REGION Network 145
   Label( C76_Comm_Fault )
   RUNG wire#powerrail
      Coil( "SectionComment" )
   END_RUNG
   // the same network as SCL:
   C76_Comm_Fault:
   "SectionComment" := TRUE;
END_REGION

REGION Network 146
   // **********************************************************************************************************************
   // 
   // Carrier 77 I-Device Data Transfer Interlocks from Carrier to SDC
   // 
   // **********************************************************************************************************************
   RUNG wire#powerrail
      Coil( "SectionComment" )
   END_RUNG
   // the same network as SCL:
   "SectionComment" := TRUE;
END_REGION

REGION Network 147
   RUNG wire#powerrail
      Contact( "Carrier_77_Status.0" )
      Coil( "EMS".Carrier[77].SDC_IN.HeartBeat )
   END_RUNG
   // the same network as SCL:
   "EMS".Carrier[77].SDC_IN.HeartBeat := "Carrier_77_Status.0";
END_REGION

REGION Network 148
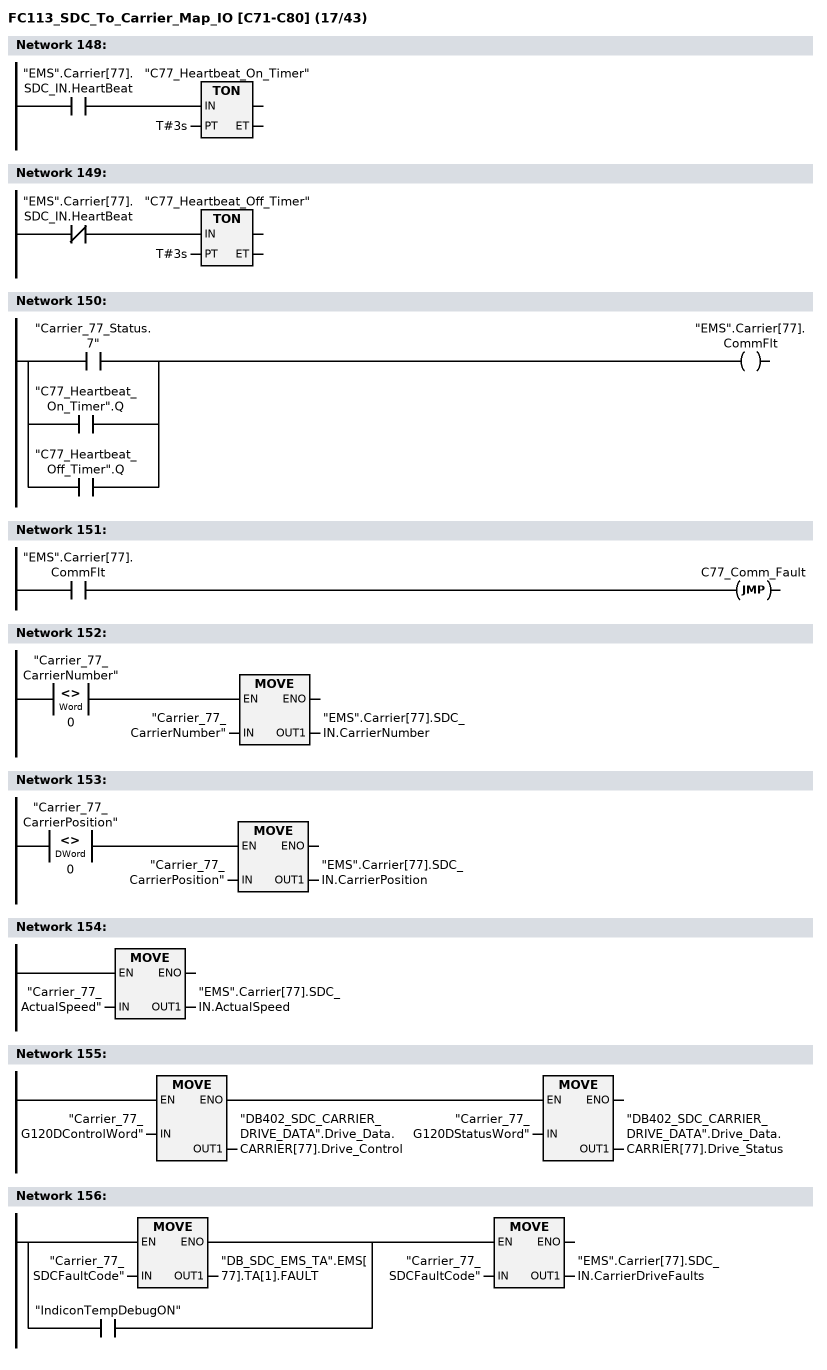
   "C77_Heartbeat_On_Timer".TON(IN := "EMS".Carrier[77].SDC_IN.HeartBeat, PT := T#3s);
END_REGION

REGION Network 149
   "C77_Heartbeat_Off_Timer".TON(IN := NOT "EMS".Carrier[77].SDC_IN.HeartBeat, PT := T#3s);
END_REGION

REGION Network 150
   RUNG wire#powerrail
      Contact( "Carrier_77_Status.7" )
      wire#w1
      Coil( "EMS".Carrier[77].CommFlt )
   END_RUNG
   RUNG wire#powerrail
      Contact( "C77_Heartbeat_On_Timer".Q )
   END_RUNG wire#w1
   RUNG wire#powerrail
      Contact( "C77_Heartbeat_Off_Timer".Q )
   END_RUNG wire#w1
   // the same network as SCL:
   "EMS".Carrier[77].CommFlt := "Carrier_77_Status.7" OR "C77_Heartbeat_On_Timer".Q OR "C77_Heartbeat_Off_Timer".Q;
END_REGION

REGION Network 151
   RUNG wire#powerrail
      Contact( "EMS".Carrier[77].CommFlt )
      JumpCoil( C77_Comm_Fault )
   END_RUNG
   // the same network as SCL:
   IF "EMS".Carrier[77].CommFlt THEN GOTO C77_Comm_Fault; END_IF;
END_REGION

REGION Network 152
   RUNG wire#powerrail
      { S7_Templates := "SrcType := Word" } NE_Contact(in1 := "Carrier_77_CarrierNumber", in2 := 0)
      Move(in := "Carrier_77_CarrierNumber", out1 => "EMS".Carrier[77].SDC_IN.CarrierNumber)
   END_RUNG
   // the same network as SCL:
   IF "Carrier_77_CarrierNumber" <> 0 THEN
       "EMS".Carrier[77].SDC_IN.CarrierNumber := "Carrier_77_CarrierNumber";
   END_IF;
END_REGION

REGION Network 153
   RUNG wire#powerrail
      { S7_Templates := "SrcType := DWord" } NE_Contact(in1 := "Carrier_77_CarrierPosition", in2 := 0)
      Move(in := "Carrier_77_CarrierPosition", out1 => "EMS".Carrier[77].SDC_IN.CarrierPosition)
   END_RUNG
   // the same network as SCL:
   IF "Carrier_77_CarrierPosition" <> 0 THEN
       "EMS".Carrier[77].SDC_IN.CarrierPosition := "Carrier_77_CarrierPosition";
   END_IF;
END_REGION

REGION Network 154
   RUNG wire#powerrail
      Move(in := "Carrier_77_ActualSpeed", out1 => "EMS".Carrier[77].SDC_IN.ActualSpeed)
   END_RUNG
   // the same network as SCL:
   "EMS".Carrier[77].SDC_IN.ActualSpeed := "Carrier_77_ActualSpeed";
END_REGION

REGION Network 155
   RUNG wire#powerrail
      Move(in := "Carrier_77_G120DControlWord", out1 => "DB402_SDC_CARRIER_DRIVE_DATA".Drive_Data.CARRIER[77].Drive_Control)
      Move(in := "Carrier_77_G120DStatusWord", out1 => "DB402_SDC_CARRIER_DRIVE_DATA".Drive_Data.CARRIER[77].Drive_Status)
   END_RUNG
   // the same network as SCL:
   "DB402_SDC_CARRIER_DRIVE_DATA".Drive_Data.CARRIER[77].Drive_Control := "Carrier_77_G120DControlWord";
   "DB402_SDC_CARRIER_DRIVE_DATA".Drive_Data.CARRIER[77].Drive_Status := "Carrier_77_G120DStatusWord";
END_REGION

REGION Network 156
   RUNG wire#powerrail
      Move(in := "Carrier_77_SDCFaultCode", out1 => "DB_SDC_EMS_TA".EMS[77].TA[1].FAULT)
      wire#w1
      Move(in := "Carrier_77_SDCFaultCode", out1 => "EMS".Carrier[77].SDC_IN.CarrierDriveFaults)
   END_RUNG
   RUNG wire#powerrail
      Contact( "IndiconTempDebugON" )
   END_RUNG wire#w1
   // the same network as SCL:
   "DB_SDC_EMS_TA".EMS[77].TA[1].FAULT := "Carrier_77_SDCFaultCode";
   IF TRUE OR "IndiconTempDebugON" THEN
       "EMS".Carrier[77].SDC_IN.CarrierDriveFaults := "Carrier_77_SDCFaultCode";
   END_IF;
END_REGION

REGION Network 157
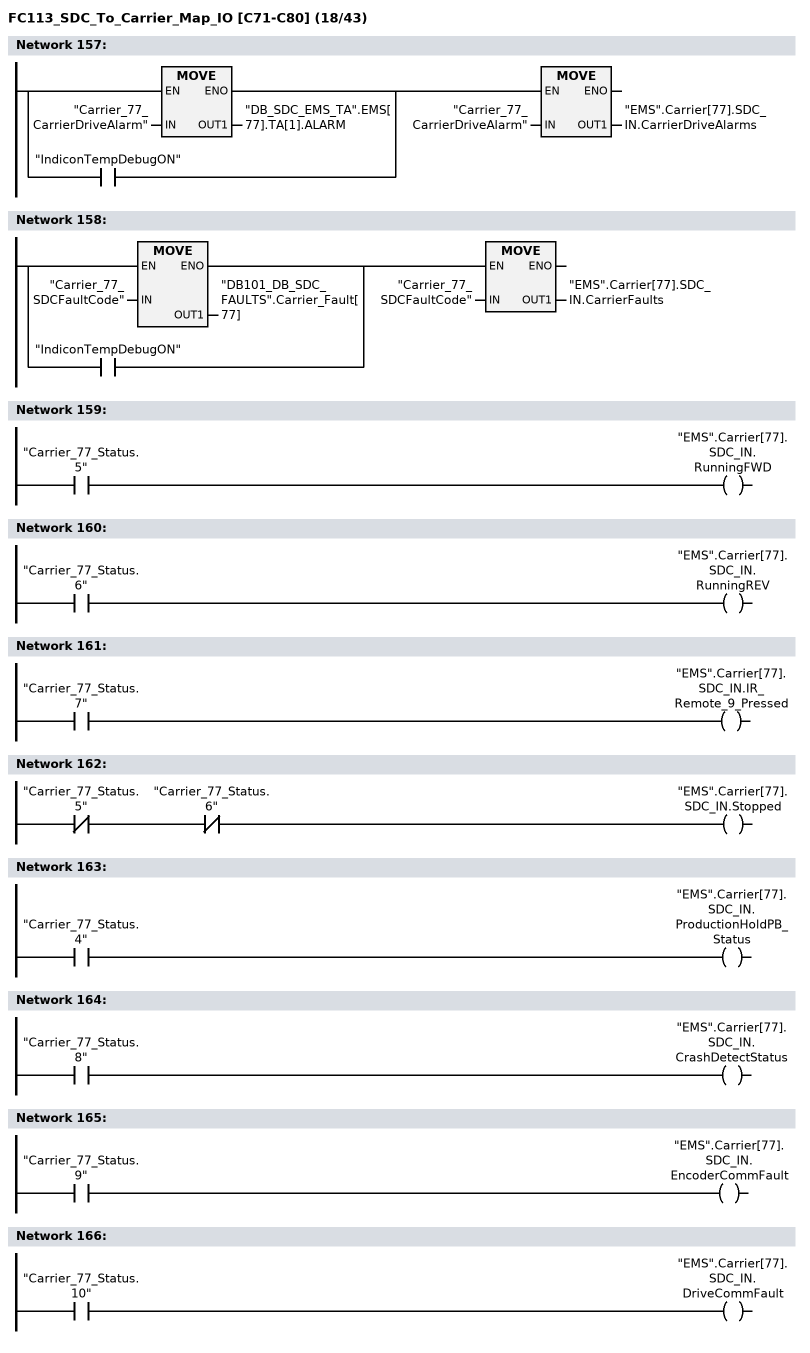
   RUNG wire#powerrail
      Move(in := "Carrier_77_CarrierDriveAlarm", out1 => "DB_SDC_EMS_TA".EMS[77].TA[1].ALARM)
      wire#w1
      Move(in := "Carrier_77_CarrierDriveAlarm", out1 => "EMS".Carrier[77].SDC_IN.CarrierDriveAlarms)
   END_RUNG
   RUNG wire#powerrail
      Contact( "IndiconTempDebugON" )
   END_RUNG wire#w1
   // the same network as SCL:
   "DB_SDC_EMS_TA".EMS[77].TA[1].ALARM := "Carrier_77_CarrierDriveAlarm";
   IF TRUE OR "IndiconTempDebugON" THEN
       "EMS".Carrier[77].SDC_IN.CarrierDriveAlarms := "Carrier_77_CarrierDriveAlarm";
   END_IF;
END_REGION

REGION Network 158
   RUNG wire#powerrail
      Move(in := "Carrier_77_SDCFaultCode", out1 => "DB101_DB_SDC_FAULTS".Carrier_Fault[77])
      wire#w1
      Move(in := "Carrier_77_SDCFaultCode", out1 => "EMS".Carrier[77].SDC_IN.CarrierFaults)
   END_RUNG
   RUNG wire#powerrail
      Contact( "IndiconTempDebugON" )
   END_RUNG wire#w1
   // the same network as SCL:
   "DB101_DB_SDC_FAULTS".Carrier_Fault[77] := "Carrier_77_SDCFaultCode";
   IF TRUE OR "IndiconTempDebugON" THEN
       "EMS".Carrier[77].SDC_IN.CarrierFaults := "Carrier_77_SDCFaultCode";
   END_IF;
END_REGION

REGION Network 159
   RUNG wire#powerrail
      Contact( "Carrier_77_Status.5" )
      Coil( "EMS".Carrier[77].SDC_IN.RunningFWD )
   END_RUNG
   // the same network as SCL:
   "EMS".Carrier[77].SDC_IN.RunningFWD := "Carrier_77_Status.5";
END_REGION

REGION Network 160
   RUNG wire#powerrail
      Contact( "Carrier_77_Status.6" )
      Coil( "EMS".Carrier[77].SDC_IN.RunningREV )
   END_RUNG
   // the same network as SCL:
   "EMS".Carrier[77].SDC_IN.RunningREV := "Carrier_77_Status.6";
END_REGION

REGION Network 161
   RUNG wire#powerrail
      Contact( "Carrier_77_Status.7" )
      Coil( "EMS".Carrier[77].SDC_IN.IR_Remote_9_Pressed )
   END_RUNG
   // the same network as SCL:
   "EMS".Carrier[77].SDC_IN.IR_Remote_9_Pressed := "Carrier_77_Status.7";
END_REGION

REGION Network 162
   RUNG wire#powerrail
      I_Contact( "Carrier_77_Status.5" )
      I_Contact( "Carrier_77_Status.6" )
      Coil( "EMS".Carrier[77].SDC_IN.Stopped )
   END_RUNG
   // the same network as SCL:
   "EMS".Carrier[77].SDC_IN.Stopped := NOT "Carrier_77_Status.5" AND NOT "Carrier_77_Status.6";
END_REGION

REGION Network 163
   RUNG wire#powerrail
      Contact( "Carrier_77_Status.4" )
      Coil( "EMS".Carrier[77].SDC_IN.ProductionHoldPB_Status )
   END_RUNG
   // the same network as SCL:
   "EMS".Carrier[77].SDC_IN.ProductionHoldPB_Status := "Carrier_77_Status.4";
END_REGION

REGION Network 164
   RUNG wire#powerrail
      Contact( "Carrier_77_Status.8" )
      Coil( "EMS".Carrier[77].SDC_IN.CrashDetectStatus )
   END_RUNG
   // the same network as SCL:
   "EMS".Carrier[77].SDC_IN.CrashDetectStatus := "Carrier_77_Status.8";
END_REGION

REGION Network 165
   RUNG wire#powerrail
      Contact( "Carrier_77_Status.9" )
      Coil( "EMS".Carrier[77].SDC_IN.EncoderCommFault )
   END_RUNG
   // the same network as SCL:
   "EMS".Carrier[77].SDC_IN.EncoderCommFault := "Carrier_77_Status.9";
END_REGION

REGION Network 166
   RUNG wire#powerrail
      Contact( "Carrier_77_Status.10" )
      Coil( "EMS".Carrier[77].SDC_IN.DriveCommFault )
   END_RUNG
   // the same network as SCL:
   "EMS".Carrier[77].SDC_IN.DriveCommFault := "Carrier_77_Status.10";
END_REGION

REGION Network 167
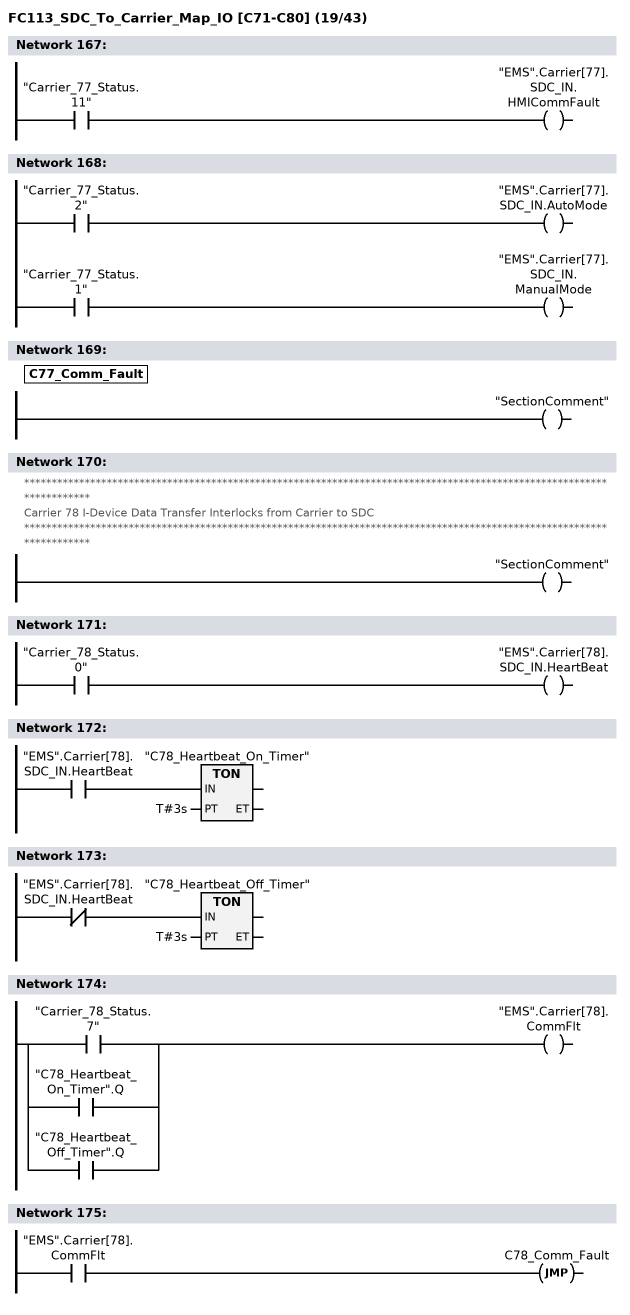
   RUNG wire#powerrail
      Contact( "Carrier_77_Status.11" )
      Coil( "EMS".Carrier[77].SDC_IN.HMICommFault )
   END_RUNG
   // the same network as SCL:
   "EMS".Carrier[77].SDC_IN.HMICommFault := "Carrier_77_Status.11";
END_REGION

REGION Network 168
   RUNG wire#powerrail
      Contact( "Carrier_77_Status.2" )
      Coil( "EMS".Carrier[77].SDC_IN.AutoMode )
   END_RUNG
   RUNG wire#powerrail
      Contact( "Carrier_77_Status.1" )
      Coil( "EMS".Carrier[77].SDC_IN.ManualMode )
   END_RUNG
   // the same network as SCL:
   "EMS".Carrier[77].SDC_IN.AutoMode := "Carrier_77_Status.2";
   "EMS".Carrier[77].SDC_IN.ManualMode := "Carrier_77_Status.1";
END_REGION

REGION Network 169
   Label( C77_Comm_Fault )
   RUNG wire#powerrail
      Coil( "SectionComment" )
   END_RUNG
   // the same network as SCL:
   C77_Comm_Fault:
   "SectionComment" := TRUE;
END_REGION

REGION Network 170
   // **********************************************************************************************************************
   // 
   // Carrier 78 I-Device Data Transfer Interlocks from Carrier to SDC
   // 
   // **********************************************************************************************************************
   RUNG wire#powerrail
      Coil( "SectionComment" )
   END_RUNG
   // the same network as SCL:
   "SectionComment" := TRUE;
END_REGION

REGION Network 171
   RUNG wire#powerrail
      Contact( "Carrier_78_Status.0" )
      Coil( "EMS".Carrier[78].SDC_IN.HeartBeat )
   END_RUNG
   // the same network as SCL:
   "EMS".Carrier[78].SDC_IN.HeartBeat := "Carrier_78_Status.0";
END_REGION

REGION Network 172
   "C78_Heartbeat_On_Timer".TON(IN := "EMS".Carrier[78].SDC_IN.HeartBeat, PT := T#3s);
END_REGION

REGION Network 173
   "C78_Heartbeat_Off_Timer".TON(IN := NOT "EMS".Carrier[78].SDC_IN.HeartBeat, PT := T#3s);
END_REGION

REGION Network 174
   RUNG wire#powerrail
      Contact( "Carrier_78_Status.7" )
      wire#w1
      Coil( "EMS".Carrier[78].CommFlt )
   END_RUNG
   RUNG wire#powerrail
      Contact( "C78_Heartbeat_On_Timer".Q )
   END_RUNG wire#w1
   RUNG wire#powerrail
      Contact( "C78_Heartbeat_Off_Timer".Q )
   END_RUNG wire#w1
   // the same network as SCL:
   "EMS".Carrier[78].CommFlt := "Carrier_78_Status.7" OR "C78_Heartbeat_On_Timer".Q OR "C78_Heartbeat_Off_Timer".Q;
END_REGION

REGION Network 175
   RUNG wire#powerrail
      Contact( "EMS".Carrier[78].CommFlt )
      JumpCoil( C78_Comm_Fault )
   END_RUNG
   // the same network as SCL:
   IF "EMS".Carrier[78].CommFlt THEN GOTO C78_Comm_Fault; END_IF;
END_REGION

REGION Network 176
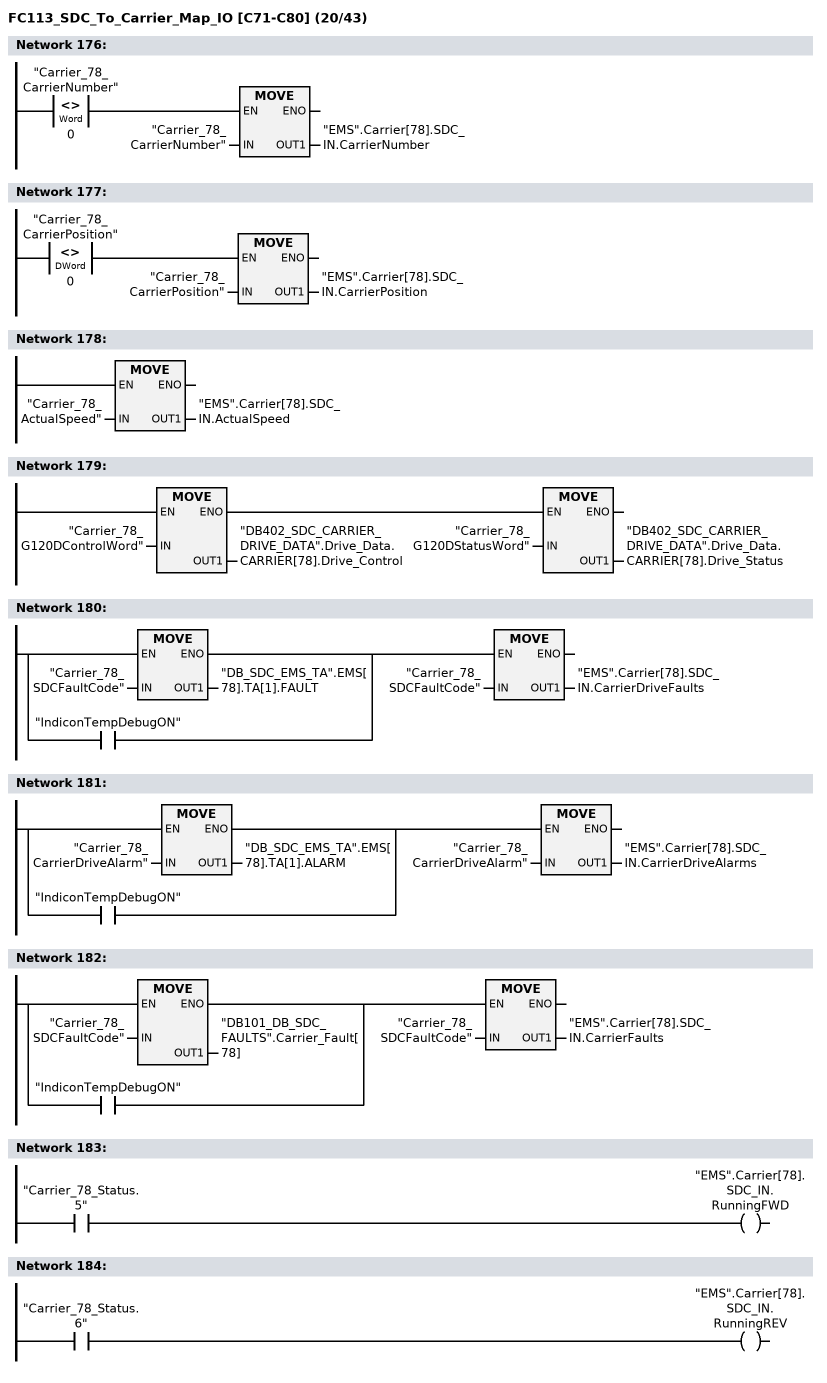
   RUNG wire#powerrail
      { S7_Templates := "SrcType := Word" } NE_Contact(in1 := "Carrier_78_CarrierNumber", in2 := 0)
      Move(in := "Carrier_78_CarrierNumber", out1 => "EMS".Carrier[78].SDC_IN.CarrierNumber)
   END_RUNG
   // the same network as SCL:
   IF "Carrier_78_CarrierNumber" <> 0 THEN
       "EMS".Carrier[78].SDC_IN.CarrierNumber := "Carrier_78_CarrierNumber";
   END_IF;
END_REGION

REGION Network 177
   RUNG wire#powerrail
      { S7_Templates := "SrcType := DWord" } NE_Contact(in1 := "Carrier_78_CarrierPosition", in2 := 0)
      Move(in := "Carrier_78_CarrierPosition", out1 => "EMS".Carrier[78].SDC_IN.CarrierPosition)
   END_RUNG
   // the same network as SCL:
   IF "Carrier_78_CarrierPosition" <> 0 THEN
       "EMS".Carrier[78].SDC_IN.CarrierPosition := "Carrier_78_CarrierPosition";
   END_IF;
END_REGION

REGION Network 178
   RUNG wire#powerrail
      Move(in := "Carrier_78_ActualSpeed", out1 => "EMS".Carrier[78].SDC_IN.ActualSpeed)
   END_RUNG
   // the same network as SCL:
   "EMS".Carrier[78].SDC_IN.ActualSpeed := "Carrier_78_ActualSpeed";
END_REGION

REGION Network 179
   RUNG wire#powerrail
      Move(in := "Carrier_78_G120DControlWord", out1 => "DB402_SDC_CARRIER_DRIVE_DATA".Drive_Data.CARRIER[78].Drive_Control)
      Move(in := "Carrier_78_G120DStatusWord", out1 => "DB402_SDC_CARRIER_DRIVE_DATA".Drive_Data.CARRIER[78].Drive_Status)
   END_RUNG
   // the same network as SCL:
   "DB402_SDC_CARRIER_DRIVE_DATA".Drive_Data.CARRIER[78].Drive_Control := "Carrier_78_G120DControlWord";
   "DB402_SDC_CARRIER_DRIVE_DATA".Drive_Data.CARRIER[78].Drive_Status := "Carrier_78_G120DStatusWord";
END_REGION

REGION Network 180
   RUNG wire#powerrail
      Move(in := "Carrier_78_SDCFaultCode", out1 => "DB_SDC_EMS_TA".EMS[78].TA[1].FAULT)
      wire#w1
      Move(in := "Carrier_78_SDCFaultCode", out1 => "EMS".Carrier[78].SDC_IN.CarrierDriveFaults)
   END_RUNG
   RUNG wire#powerrail
      Contact( "IndiconTempDebugON" )
   END_RUNG wire#w1
   // the same network as SCL:
   "DB_SDC_EMS_TA".EMS[78].TA[1].FAULT := "Carrier_78_SDCFaultCode";
   IF TRUE OR "IndiconTempDebugON" THEN
       "EMS".Carrier[78].SDC_IN.CarrierDriveFaults := "Carrier_78_SDCFaultCode";
   END_IF;
END_REGION

REGION Network 181
   RUNG wire#powerrail
      Move(in := "Carrier_78_CarrierDriveAlarm", out1 => "DB_SDC_EMS_TA".EMS[78].TA[1].ALARM)
      wire#w1
      Move(in := "Carrier_78_CarrierDriveAlarm", out1 => "EMS".Carrier[78].SDC_IN.CarrierDriveAlarms)
   END_RUNG
   RUNG wire#powerrail
      Contact( "IndiconTempDebugON" )
   END_RUNG wire#w1
   // the same network as SCL:
   "DB_SDC_EMS_TA".EMS[78].TA[1].ALARM := "Carrier_78_CarrierDriveAlarm";
   IF TRUE OR "IndiconTempDebugON" THEN
       "EMS".Carrier[78].SDC_IN.CarrierDriveAlarms := "Carrier_78_CarrierDriveAlarm";
   END_IF;
END_REGION

REGION Network 182
   RUNG wire#powerrail
      Move(in := "Carrier_78_SDCFaultCode", out1 => "DB101_DB_SDC_FAULTS".Carrier_Fault[78])
      wire#w1
      Move(in := "Carrier_78_SDCFaultCode", out1 => "EMS".Carrier[78].SDC_IN.CarrierFaults)
   END_RUNG
   RUNG wire#powerrail
      Contact( "IndiconTempDebugON" )
   END_RUNG wire#w1
   // the same network as SCL:
   "DB101_DB_SDC_FAULTS".Carrier_Fault[78] := "Carrier_78_SDCFaultCode";
   IF TRUE OR "IndiconTempDebugON" THEN
       "EMS".Carrier[78].SDC_IN.CarrierFaults := "Carrier_78_SDCFaultCode";
   END_IF;
END_REGION

REGION Network 183
   RUNG wire#powerrail
      Contact( "Carrier_78_Status.5" )
      Coil( "EMS".Carrier[78].SDC_IN.RunningFWD )
   END_RUNG
   // the same network as SCL:
   "EMS".Carrier[78].SDC_IN.RunningFWD := "Carrier_78_Status.5";
END_REGION

REGION Network 184
   RUNG wire#powerrail
      Contact( "Carrier_78_Status.6" )
      Coil( "EMS".Carrier[78].SDC_IN.RunningREV )
   END_RUNG
   // the same network as SCL:
   "EMS".Carrier[78].SDC_IN.RunningREV := "Carrier_78_Status.6";
END_REGION

REGION Network 185
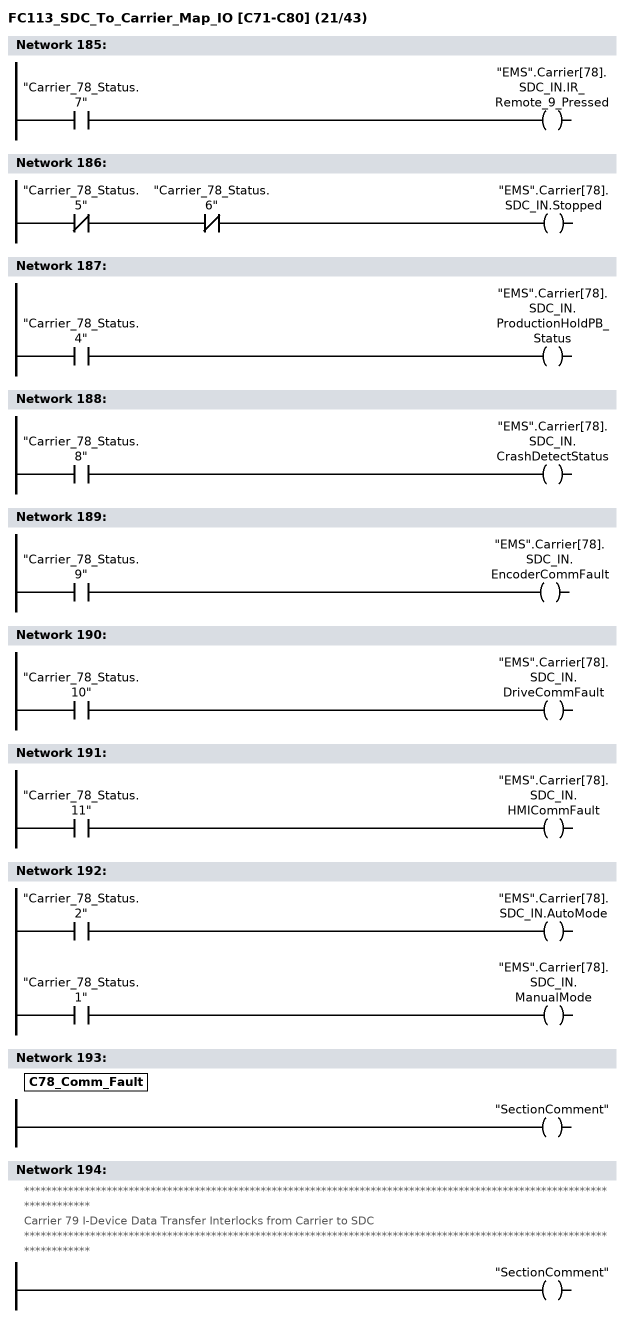
   RUNG wire#powerrail
      Contact( "Carrier_78_Status.7" )
      Coil( "EMS".Carrier[78].SDC_IN.IR_Remote_9_Pressed )
   END_RUNG
   // the same network as SCL:
   "EMS".Carrier[78].SDC_IN.IR_Remote_9_Pressed := "Carrier_78_Status.7";
END_REGION

REGION Network 186
   RUNG wire#powerrail
      I_Contact( "Carrier_78_Status.5" )
      I_Contact( "Carrier_78_Status.6" )
      Coil( "EMS".Carrier[78].SDC_IN.Stopped )
   END_RUNG
   // the same network as SCL:
   "EMS".Carrier[78].SDC_IN.Stopped := NOT "Carrier_78_Status.5" AND NOT "Carrier_78_Status.6";
END_REGION

REGION Network 187
   RUNG wire#powerrail
      Contact( "Carrier_78_Status.4" )
      Coil( "EMS".Carrier[78].SDC_IN.ProductionHoldPB_Status )
   END_RUNG
   // the same network as SCL:
   "EMS".Carrier[78].SDC_IN.ProductionHoldPB_Status := "Carrier_78_Status.4";
END_REGION

REGION Network 188
   RUNG wire#powerrail
      Contact( "Carrier_78_Status.8" )
      Coil( "EMS".Carrier[78].SDC_IN.CrashDetectStatus )
   END_RUNG
   // the same network as SCL:
   "EMS".Carrier[78].SDC_IN.CrashDetectStatus := "Carrier_78_Status.8";
END_REGION

REGION Network 189
   RUNG wire#powerrail
      Contact( "Carrier_78_Status.9" )
      Coil( "EMS".Carrier[78].SDC_IN.EncoderCommFault )
   END_RUNG
   // the same network as SCL:
   "EMS".Carrier[78].SDC_IN.EncoderCommFault := "Carrier_78_Status.9";
END_REGION

REGION Network 190
   RUNG wire#powerrail
      Contact( "Carrier_78_Status.10" )
      Coil( "EMS".Carrier[78].SDC_IN.DriveCommFault )
   END_RUNG
   // the same network as SCL:
   "EMS".Carrier[78].SDC_IN.DriveCommFault := "Carrier_78_Status.10";
END_REGION

REGION Network 191
   RUNG wire#powerrail
      Contact( "Carrier_78_Status.11" )
      Coil( "EMS".Carrier[78].SDC_IN.HMICommFault )
   END_RUNG
   // the same network as SCL:
   "EMS".Carrier[78].SDC_IN.HMICommFault := "Carrier_78_Status.11";
END_REGION

REGION Network 192
   RUNG wire#powerrail
      Contact( "Carrier_78_Status.2" )
      Coil( "EMS".Carrier[78].SDC_IN.AutoMode )
   END_RUNG
   RUNG wire#powerrail
      Contact( "Carrier_78_Status.1" )
      Coil( "EMS".Carrier[78].SDC_IN.ManualMode )
   END_RUNG
   // the same network as SCL:
   "EMS".Carrier[78].SDC_IN.AutoMode := "Carrier_78_Status.2";
   "EMS".Carrier[78].SDC_IN.ManualMode := "Carrier_78_Status.1";
END_REGION

REGION Network 193
   Label( C78_Comm_Fault )
   RUNG wire#powerrail
      Coil( "SectionComment" )
   END_RUNG
   // the same network as SCL:
   C78_Comm_Fault:
   "SectionComment" := TRUE;
END_REGION

REGION Network 194
   // **********************************************************************************************************************
   // 
   // Carrier 79 I-Device Data Transfer Interlocks from Carrier to SDC
   // 
   // **********************************************************************************************************************
   RUNG wire#powerrail
      Coil( "SectionComment" )
   END_RUNG
   // the same network as SCL:
   "SectionComment" := TRUE;
END_REGION

REGION Network 195
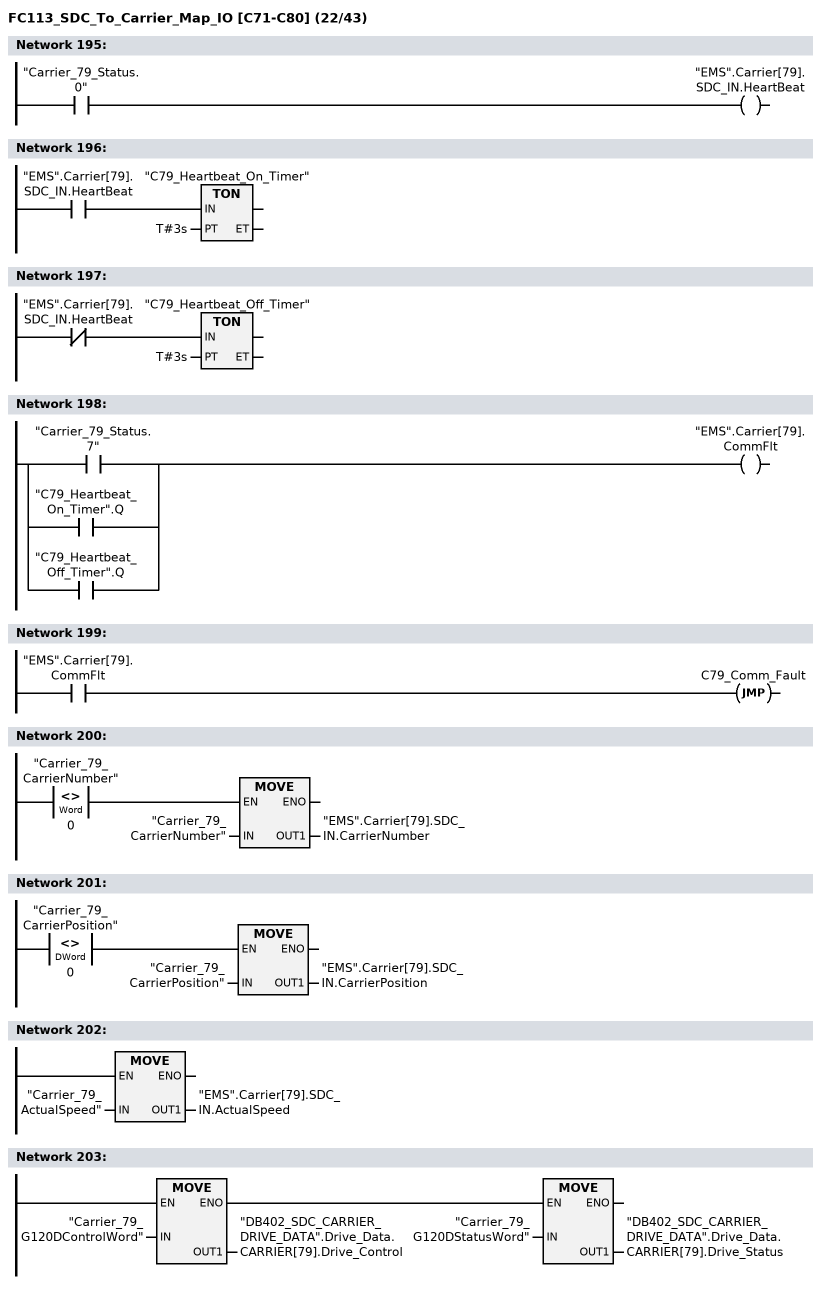
   RUNG wire#powerrail
      Contact( "Carrier_79_Status.0" )
      Coil( "EMS".Carrier[79].SDC_IN.HeartBeat )
   END_RUNG
   // the same network as SCL:
   "EMS".Carrier[79].SDC_IN.HeartBeat := "Carrier_79_Status.0";
END_REGION

REGION Network 196
   "C79_Heartbeat_On_Timer".TON(IN := "EMS".Carrier[79].SDC_IN.HeartBeat, PT := T#3s);
END_REGION

REGION Network 197
   "C79_Heartbeat_Off_Timer".TON(IN := NOT "EMS".Carrier[79].SDC_IN.HeartBeat, PT := T#3s);
END_REGION

REGION Network 198
   RUNG wire#powerrail
      Contact( "Carrier_79_Status.7" )
      wire#w1
      Coil( "EMS".Carrier[79].CommFlt )
   END_RUNG
   RUNG wire#powerrail
      Contact( "C79_Heartbeat_On_Timer".Q )
   END_RUNG wire#w1
   RUNG wire#powerrail
      Contact( "C79_Heartbeat_Off_Timer".Q )
   END_RUNG wire#w1
   // the same network as SCL:
   "EMS".Carrier[79].CommFlt := "Carrier_79_Status.7" OR "C79_Heartbeat_On_Timer".Q OR "C79_Heartbeat_Off_Timer".Q;
END_REGION

REGION Network 199
   RUNG wire#powerrail
      Contact( "EMS".Carrier[79].CommFlt )
      JumpCoil( C79_Comm_Fault )
   END_RUNG
   // the same network as SCL:
   IF "EMS".Carrier[79].CommFlt THEN GOTO C79_Comm_Fault; END_IF;
END_REGION

REGION Network 200
   RUNG wire#powerrail
      { S7_Templates := "SrcType := Word" } NE_Contact(in1 := "Carrier_79_CarrierNumber", in2 := 0)
      Move(in := "Carrier_79_CarrierNumber", out1 => "EMS".Carrier[79].SDC_IN.CarrierNumber)
   END_RUNG
   // the same network as SCL:
   IF "Carrier_79_CarrierNumber" <> 0 THEN
       "EMS".Carrier[79].SDC_IN.CarrierNumber := "Carrier_79_CarrierNumber";
   END_IF;
END_REGION

REGION Network 201
   RUNG wire#powerrail
      { S7_Templates := "SrcType := DWord" } NE_Contact(in1 := "Carrier_79_CarrierPosition", in2 := 0)
      Move(in := "Carrier_79_CarrierPosition", out1 => "EMS".Carrier[79].SDC_IN.CarrierPosition)
   END_RUNG
   // the same network as SCL:
   IF "Carrier_79_CarrierPosition" <> 0 THEN
       "EMS".Carrier[79].SDC_IN.CarrierPosition := "Carrier_79_CarrierPosition";
   END_IF;
END_REGION

REGION Network 202
   RUNG wire#powerrail
      Move(in := "Carrier_79_ActualSpeed", out1 => "EMS".Carrier[79].SDC_IN.ActualSpeed)
   END_RUNG
   // the same network as SCL:
   "EMS".Carrier[79].SDC_IN.ActualSpeed := "Carrier_79_ActualSpeed";
END_REGION

REGION Network 203
   RUNG wire#powerrail
      Move(in := "Carrier_79_G120DControlWord", out1 => "DB402_SDC_CARRIER_DRIVE_DATA".Drive_Data.CARRIER[79].Drive_Control)
      Move(in := "Carrier_79_G120DStatusWord", out1 => "DB402_SDC_CARRIER_DRIVE_DATA".Drive_Data.CARRIER[79].Drive_Status)
   END_RUNG
   // the same network as SCL:
   "DB402_SDC_CARRIER_DRIVE_DATA".Drive_Data.CARRIER[79].Drive_Control := "Carrier_79_G120DControlWord";
   "DB402_SDC_CARRIER_DRIVE_DATA".Drive_Data.CARRIER[79].Drive_Status := "Carrier_79_G120DStatusWord";
END_REGION

REGION Network 204
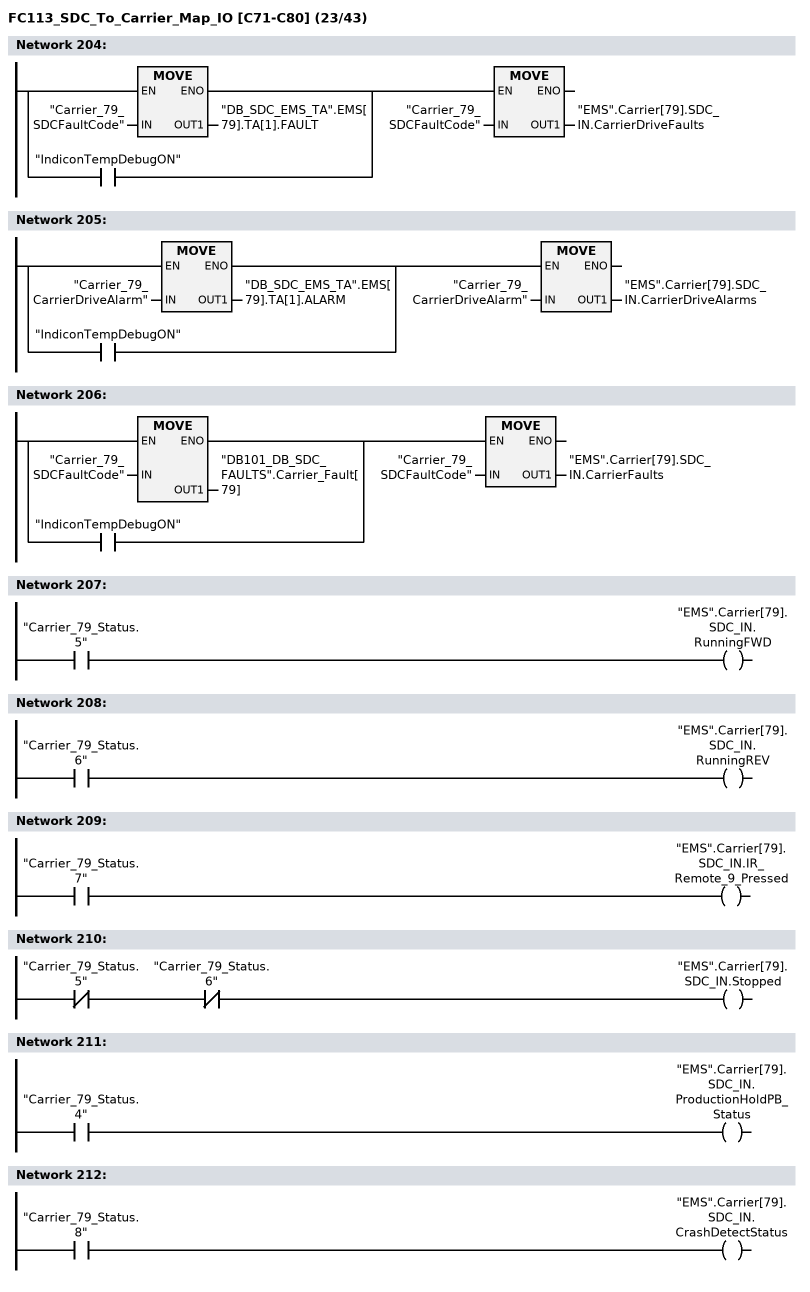
   RUNG wire#powerrail
      Move(in := "Carrier_79_SDCFaultCode", out1 => "DB_SDC_EMS_TA".EMS[79].TA[1].FAULT)
      wire#w1
      Move(in := "Carrier_79_SDCFaultCode", out1 => "EMS".Carrier[79].SDC_IN.CarrierDriveFaults)
   END_RUNG
   RUNG wire#powerrail
      Contact( "IndiconTempDebugON" )
   END_RUNG wire#w1
   // the same network as SCL:
   "DB_SDC_EMS_TA".EMS[79].TA[1].FAULT := "Carrier_79_SDCFaultCode";
   IF TRUE OR "IndiconTempDebugON" THEN
       "EMS".Carrier[79].SDC_IN.CarrierDriveFaults := "Carrier_79_SDCFaultCode";
   END_IF;
END_REGION

REGION Network 205
   RUNG wire#powerrail
      Move(in := "Carrier_79_CarrierDriveAlarm", out1 => "DB_SDC_EMS_TA".EMS[79].TA[1].ALARM)
      wire#w1
      Move(in := "Carrier_79_CarrierDriveAlarm", out1 => "EMS".Carrier[79].SDC_IN.CarrierDriveAlarms)
   END_RUNG
   RUNG wire#powerrail
      Contact( "IndiconTempDebugON" )
   END_RUNG wire#w1
   // the same network as SCL:
   "DB_SDC_EMS_TA".EMS[79].TA[1].ALARM := "Carrier_79_CarrierDriveAlarm";
   IF TRUE OR "IndiconTempDebugON" THEN
       "EMS".Carrier[79].SDC_IN.CarrierDriveAlarms := "Carrier_79_CarrierDriveAlarm";
   END_IF;
END_REGION

REGION Network 206
   RUNG wire#powerrail
      Move(in := "Carrier_79_SDCFaultCode", out1 => "DB101_DB_SDC_FAULTS".Carrier_Fault[79])
      wire#w1
      Move(in := "Carrier_79_SDCFaultCode", out1 => "EMS".Carrier[79].SDC_IN.CarrierFaults)
   END_RUNG
   RUNG wire#powerrail
      Contact( "IndiconTempDebugON" )
   END_RUNG wire#w1
   // the same network as SCL:
   "DB101_DB_SDC_FAULTS".Carrier_Fault[79] := "Carrier_79_SDCFaultCode";
   IF TRUE OR "IndiconTempDebugON" THEN
       "EMS".Carrier[79].SDC_IN.CarrierFaults := "Carrier_79_SDCFaultCode";
   END_IF;
END_REGION

REGION Network 207
   RUNG wire#powerrail
      Contact( "Carrier_79_Status.5" )
      Coil( "EMS".Carrier[79].SDC_IN.RunningFWD )
   END_RUNG
   // the same network as SCL:
   "EMS".Carrier[79].SDC_IN.RunningFWD := "Carrier_79_Status.5";
END_REGION

REGION Network 208
   RUNG wire#powerrail
      Contact( "Carrier_79_Status.6" )
      Coil( "EMS".Carrier[79].SDC_IN.RunningREV )
   END_RUNG
   // the same network as SCL:
   "EMS".Carrier[79].SDC_IN.RunningREV := "Carrier_79_Status.6";
END_REGION

REGION Network 209
   RUNG wire#powerrail
      Contact( "Carrier_79_Status.7" )
      Coil( "EMS".Carrier[79].SDC_IN.IR_Remote_9_Pressed )
   END_RUNG
   // the same network as SCL:
   "EMS".Carrier[79].SDC_IN.IR_Remote_9_Pressed := "Carrier_79_Status.7";
END_REGION

REGION Network 210
   RUNG wire#powerrail
      I_Contact( "Carrier_79_Status.5" )
      I_Contact( "Carrier_79_Status.6" )
      Coil( "EMS".Carrier[79].SDC_IN.Stopped )
   END_RUNG
   // the same network as SCL:
   "EMS".Carrier[79].SDC_IN.Stopped := NOT "Carrier_79_Status.5" AND NOT "Carrier_79_Status.6";
END_REGION

REGION Network 211
   RUNG wire#powerrail
      Contact( "Carrier_79_Status.4" )
      Coil( "EMS".Carrier[79].SDC_IN.ProductionHoldPB_Status )
   END_RUNG
   // the same network as SCL:
   "EMS".Carrier[79].SDC_IN.ProductionHoldPB_Status := "Carrier_79_Status.4";
END_REGION

REGION Network 212
   RUNG wire#powerrail
      Contact( "Carrier_79_Status.8" )
      Coil( "EMS".Carrier[79].SDC_IN.CrashDetectStatus )
   END_RUNG
   // the same network as SCL:
   "EMS".Carrier[79].SDC_IN.CrashDetectStatus := "Carrier_79_Status.8";
END_REGION

REGION Network 213